
Template "Navigation" 1280x800
   TextField "Template_Text field_1" at 1044,28 size 229x39; Text 'Krauss Maffei'
   Button "Template_Button_17" at 502,23 size 38x32; TextOff 'Text'; PictureOff "Bendera inggris"
      on Click: function_fb9197e8(-1)
   Button "Template_Button_18" at 546,23 size 38x32; TextOff 'Text'; PictureOff "manual mode"
   Button "Template_Button_19" at 590,23 size 38x32; TextOff 'Text'; PictureOff "automatic mode"; PictureList "Operation Mode"
      ProcessValue <- "Operation Mode"
   Button "Template_Button_20" at 634,23 size 38x32; TextOff 'Text'
   Button "Template_Button_21" at 678,23 size 38x32; TextOff 'Text'
   Button "Template_Button_24" at 16,18 size 67x43; TextOff 'Text'; PictureOff "left arrow"
      on Press: function_efd93a16()
   Button "status_reduced" at 678,23 size 38x32; TextOff 'Text'; PictureOff "Reduced green"
      Visibility <- "DB619_State_MPart_Recirculation{1}_Reduced"
   Button "Template_Button_15" at 414,23 size 38x32; TextOff 'Text'
   Button "status_Interval_Reduced" at 678,23 size 38x32; TextOff 'Text'; PictureOff "Interval green"
      Visibility <- "DB619_State_MPart_Recirculation{1}_Intervall_Reduced"
   Button "status_lowpressure" at 678,23 size 38x32; TextOff 'Text'; PictureOff "Lowpress green"
      Visibility <- "DB619_State_MPart_Recirculation{1}_Lowpressure"
   Button "status_Lowpressure_Interval" at 678,23 size 38x32; TextOff 'Text'; PictureOff "lowpress circulation"
      Visibility <- "DB619_State_MPart_Recirculation{1}_Intervall_Lowpressure"
   Button "status_highpressure" at 678,23 size 38x32; TextOff 'Text'; PictureOff "high press circuit"
      Visibility <- "DB619_State_MPart_Recirculation{1}_Highpressure"
   Button "Template_Button_25" at 546,23 size 38x32; TextOff 'Text'; PictureList "Operation Mode"; PictureOff "weekendmode"
      ProcessValue <- "Operation Mode"
      Visibility <- "DB619_State_MPart_Recirculation{1}_Weekendswitching"
   Button "Template_Button_26" at 722,23 size 38x32; TextOff 'Text'
   Button "Template_Button_27" at 678,23 size 38x32; TextOff 'Text'; PictureOff "shot cycle_1"
      Visibility <- "DB619_State_MPart_Cycle{1}_running"
   IOField "Template_I/O field_1" at 97,25 size 273x28; FormatPattern 9999999999999999999999999999999999999999
      ProcessValue <- "TP-Bereichszeiger_Date_Time_ActTime"
   Button "Template_Button_30" at 458,23 size 38x32; TextOff 'Text'
   Button "Template_Button_16" at 458,23 size 38x32; TextOff 'Text'; PictureOff "printer off"; PictureList "Print Function"
      ProcessValue <- "Print Function"
      Visibility <- "Print Function"
   SymbolicIOField "Template_Symbolic I/O field_1" at 800,18 size 120x42; TextOff '0'; TextOn '1'; TextList "MH_NO"
      ProcessValue <- "DB619_State_MPart_SWU{1}_ActualSWU"
   Button "Template_Button_3" at 16,261 size 68x66; TextOff 'Text'; PictureOff "osiloskope"; PictureList "ico_navigation_1"
      on Press: function_b14e0dd5("DB14_TP_Shortcuts_TP_Shortcuts_ButtonNo_2", 0)
      Appearance <- "DB14_TP_Shortcuts_TP_Shortcuts_Page_active_2"
      on Click: ActivateScreenByNumber("DB14_TP_Shortcuts_TP_Shortcuts_PageNo_2", 0)
      Visibility <- "DB14_TP_Shortcuts_TP_Shortcuts_Page_active_2"
      ProcessValue <- "DB14_TP_Shortcuts_TP_Shortcuts_PageNo_2"
   Button "Template_Button_4" at 16,354 size 68x66; TextOff 'Text'; PictureOff "scope_1"; PictureList "ico_navigation_1"
      on Press: function_b14e0dd5("DB14_TP_Shortcuts_TP_Shortcuts_ButtonNo_3", 0)
      on Click: ActivateScreenByNumber("DB14_TP_Shortcuts_TP_Shortcuts_PageNo_3", 0)
      Appearance <- "DB14_TP_Shortcuts_TP_Shortcuts_Page_active_3"
      Visibility <- "DB14_TP_Shortcuts_TP_Shortcuts_Page_active_3"
      ProcessValue <- "DB14_TP_Shortcuts_TP_Shortcuts_PageNo_3"
   Button "Template_Button_6" at 16,539 size 68x66; TextOff 'Text'; PictureOff "s2"; PictureList "ico_navigation_1"
      on Press: function_b14e0dd5("DB14_TP_Shortcuts_TP_Shortcuts_ButtonNo_5", 0)
      on Click: ActivateScreenByNumber("DB14_TP_Shortcuts_TP_Shortcuts_PageNo_5", 0)
      Appearance <- "DB14_TP_Shortcuts_TP_Shortcuts_Page_active_5"
      Visibility <- "DB14_TP_Shortcuts_TP_Shortcuts_Page_active_5"
      ProcessValue <- "DB14_TP_Shortcuts_TP_Shortcuts_PageNo_5"
   Button "Template_Button_13" at 1196,724 size 68x66; TextOff 'Text'; PictureList "Home"; PictureOff "Graphic_8"
      on Click: ActivateScreen("0017_Home Screen", 0)
      Appearance <- "NavScreenChange"
   Button "Template_Button_23" at 1196,631 size 68x66; TextOff 'Text'; PictureList "Nav_Recipe"; PictureOff "chemical"
      on Click: ActivateScreen("0892_Tool Editor", 0)
      Appearance <- "NavScreenChange"
   Button "Template_Button_22" at 1196,446 size 68x66; TextOff 'Text'; PictureOff "archive"; PictureList "Nav_Logging"
      on Click: SetTag("NavScreenChange", 4); SetTag("Recipe_Appearance_Control", 0); SetTag("Archived Alarm Control", 2); SetTag("Archive Alarm Number", 0); "CopyAlarmLogView"(); ActivateScreen("0013_Archive Alarm", 0)
      Appearance <- "NavScreenChange"
   Button "Template_Button_9" at 1196,261 size 68x66; TextOff 'Text'; PictureOff "process"; PictureList "Setting"
      on Click: ActivateScreen("0018_SystemSetting", 0); SetTag("System Setting Screen Control", 0)
      Appearance <- "NavScreenChange"
   Button "Template_Button_2" at 16,169 size 68x66; TextOff 'Text'; PictureList "ico_navigation_1"
      on Press: function_b14e0dd5("DB14_TP_Shortcuts_TP_Shortcuts_ButtonNo_1", 0)
      on Click: ActivateScreenByNumber("DB14_TP_Shortcuts_TP_Shortcuts_PageNo_1", 0)
      Appearance <- "DB14_TP_Shortcuts_TP_Shortcuts_Page_active_1"
      Visibility <- "DB14_TP_Shortcuts_TP_Shortcuts_Page_active_1"
      ProcessValue <- "DB14_TP_Shortcuts_TP_Shortcuts_PageNo_1"
   Button "Template_Button_5" at 16,446 size 68x66; TextOff 'Text'; PictureList "ico_navigation_1"
      on Press: function_b14e0dd5("DB14_TP_Shortcuts_TP_Shortcuts_ButtonNo_4", 0)
      on Click: ActivateScreenByNumber("DB14_TP_Shortcuts_TP_Shortcuts_PageNo_4", 0)
      Appearance <- "DB14_TP_Shortcuts_TP_Shortcuts_Page_active_4"
      Visibility <- "DB14_TP_Shortcuts_TP_Shortcuts_Page_active_4"
      ProcessValue <- "DB14_TP_Shortcuts_TP_Shortcuts_PageNo_4"
   Button "Template_Button_31" at 16,631 size 68x66; TextOff 'Text'; PictureOff "scope_1"; PictureList "ico_navigation_1"
      on Press: function_b14e0dd5("DB14_TP_Shortcuts_TP_Shortcuts_ButtonNo_6", 0)
      on Click: ActivateScreenByNumber("DB14_TP_Shortcuts_TP_Shortcuts_PageNo_6", 0)
      Appearance <- "DB14_TP_Shortcuts_TP_Shortcuts_Page_active_6"
      Visibility <- "DB14_TP_Shortcuts_TP_Shortcuts_Page_active_6"
      ProcessValue <- "DB14_TP_Shortcuts_TP_Shortcuts_PageNo_6"
   Button "Template_Button_7" at 16,724 size 68x66; TextOff 'Text'; PictureList "ico_navigation_1"
      on Press: function_b14e0dd5("DB14_TP_Shortcuts_TP_Shortcuts_ButtonNo_7", 0)
      on Click: ActivateScreenByNumber("DB14_TP_Shortcuts_TP_Shortcuts_PageNo_7", 0)
      Appearance <- "DB14_TP_Shortcuts_TP_Shortcuts_Page_active_7"
      Visibility <- "DB14_TP_Shortcuts_TP_Shortcuts_Page_active_7"
      ProcessValue <- "DB14_TP_Shortcuts_TP_Shortcuts_PageNo_7"
   Button "Template_Button_8" at 1196,169 size 68x66; TextOff 'Text'; PictureOff "Alarm Icon 3"
      on Click: ActivateScreen("0024_ActualFaults", 0); SetTag("NavScreenChange", 1); SetTag("Recipe_Appearance_Control", 0); SetTag("Alarm_Filter_Tag", 0)
      Appearance <- "NavScreenChange"
   Button "Template_Button_10" at 1196,354 size 68x66; TextOff 'Text'
   Button "Template_Button_32" at 1196,539 size 68x66; TextOff 'Text'; PictureOff "049-book"
      on Click: ActivateScreen("0999_Service", 0); SetTag("Service Screen Control Visibility", 0)
      Appearance <- "NavScreenChange"
   Button "Template_Button_11" at 371,23 size 38x32; TextOff 'Text'
      on Click: function_a2a04561()
      Appearance <- "NavUserChange"
   Button "Template_Button_33" at 16,261 size 68x66; TextOff 'Text'; PictureOff "osiloskope"; PictureList "Ico_navigation_2"
      on Click: ActivateScreenByNumber("DB14_TP_Shortcuts_TP_Shortcuts_PageNo_2", 0)
      on Press: function_b14e0dd5("DB14_TP_Shortcuts_TP_Shortcuts_ButtonNo_2", 0)
      Appearance <- "DB14_TP_Shortcuts_TP_Shortcuts_Page_active_2"
      Visibility <- "DB14_TP_Shortcuts_TP_Shortcuts_Page_active_2"
      ProcessValue <- "DB14_TP_Shortcuts_TP_Shortcuts_PageNo_2"
   Button "Template_Button_34" at 16,354 size 68x66; TextOff 'Text'; PictureOff "scope_1"; PictureList "Ico_navigation_2"
      on Press: function_b14e0dd5("DB14_TP_Shortcuts_TP_Shortcuts_ButtonNo_3", 0)
      Appearance <- "DB14_TP_Shortcuts_TP_Shortcuts_Page_active_3"
      Visibility <- "DB14_TP_Shortcuts_TP_Shortcuts_Page_active_3"
      on Click: ActivateScreenByNumber("DB14_TP_Shortcuts_TP_Shortcuts_PageNo_3", 0)
      ProcessValue <- "DB14_TP_Shortcuts_TP_Shortcuts_PageNo_3"
   Button "Template_Button_35" at 16,539 size 68x66; TextOff 'Text'; PictureOff "s2"; PictureList "Ico_navigation_2"
      on Press: function_b14e0dd5("DB14_TP_Shortcuts_TP_Shortcuts_ButtonNo_5", 0)
      Appearance <- "DB14_TP_Shortcuts_TP_Shortcuts_Page_active_5"
      Visibility <- "DB14_TP_Shortcuts_TP_Shortcuts_Page_active_5"
      on Click: ActivateScreenByNumber("DB14_TP_Shortcuts_TP_Shortcuts_PageNo_5", 0)
      ProcessValue <- "DB14_TP_Shortcuts_TP_Shortcuts_PageNo_5"
   Button "Template_Button_36" at 16,169 size 68x66; TextOff 'Text'; PictureList "Ico_navigation_2"
      on Click: ActivateScreenByNumber("DB14_TP_Shortcuts_TP_Shortcuts_PageNo_1", 0)
      on Press: function_b14e0dd5("DB14_TP_Shortcuts_TP_Shortcuts_ButtonNo_1", 0)
      Appearance <- "DB14_TP_Shortcuts_TP_Shortcuts_Page_active_1"
      Visibility <- "DB14_TP_Shortcuts_TP_Shortcuts_Page_active_1"
      ProcessValue <- "DB14_TP_Shortcuts_TP_Shortcuts_PageNo_1"
   Button "Template_Button_37" at 16,446 size 68x66; TextOff 'Text'; PictureList "Ico_navigation_2"
      on Press: function_b14e0dd5("DB14_TP_Shortcuts_TP_Shortcuts_ButtonNo_4", 0)
      Appearance <- "DB14_TP_Shortcuts_TP_Shortcuts_Page_active_4"
      Visibility <- "DB14_TP_Shortcuts_TP_Shortcuts_Page_active_4"
      on Click: ActivateScreenByNumber("DB14_TP_Shortcuts_TP_Shortcuts_PageNo_4", 0)
      ProcessValue <- "DB14_TP_Shortcuts_TP_Shortcuts_PageNo_4"
   Button "Template_Button_38" at 16,631 size 68x66; TextOff 'Text'; PictureOff "scope_1"; PictureList "Ico_navigation_2"
      on Press: function_b14e0dd5("DB14_TP_Shortcuts_TP_Shortcuts_ButtonNo_6", 0)
      Appearance <- "DB14_TP_Shortcuts_TP_Shortcuts_Page_active_6"
      Visibility <- "DB14_TP_Shortcuts_TP_Shortcuts_Page_active_6"
      on Click: ActivateScreenByNumber("DB14_TP_Shortcuts_TP_Shortcuts_PageNo_6", 0)
      ProcessValue <- "DB14_TP_Shortcuts_TP_Shortcuts_PageNo_6"
   Button "Template_Button_39" at 16,724 size 68x66; TextOff 'Text'; PictureList "Ico_navigation_2"
      on Press: function_b14e0dd5("DB14_TP_Shortcuts_TP_Shortcuts_ButtonNo_7", 0)
      Appearance <- "DB14_TP_Shortcuts_TP_Shortcuts_Page_active_7"
      Visibility <- "DB14_TP_Shortcuts_TP_Shortcuts_Page_active_7"
      on Click: ActivateScreenByNumber("DB14_TP_Shortcuts_TP_Shortcuts_PageNo_7", 0)
      ProcessValue <- "DB14_TP_Shortcuts_TP_Shortcuts_PageNo_7"
   Button "Template_Button_40" at 9,160 size 80x636; TextOff 'Text'
      on Click: function_efd93a16("Save", 446, 387, -1, 1, 1)
      Visibility <- "DB_MouldEditor_HMI_uData_sStatusBits"
   Button "Template_Button_47" at 1189,147 size 80x645; TextOff 'Text'
      Visibility <- "DB_MouldEditor_HMI_uData_sStatusBits_xValueChanged"
      on Click: function_efd93a16("Save", 446, 387, -1, -1, 1)
   Button "Template_Button_12" at 9,160 size 80x636; TextOff 'Text'
      on Click: function_efd93a16("Save", 446, 387, -1, -1, 1)
      Visibility <- "DB_MouldEditor_HMI_uData_sStatusBits"
   Button "Template_Button_14" at 1189,147 size 80x645; TextOff 'Text'
      on Click: function_efd93a16("Save", 446, 387, -1, -1, 1)
      Visibility <- "DB_MouldEditor_HMI_uData_sStatusBits_xValueChanged"
      ObjectEnable <- "PopUp_Restrict"
   Button "Template_Button_29" at 9,147 size 80x645; TextOff 'Text'
      on Click: function_efd93a16("Save", 446, 387, -1, -1, 1)
      Visibility <- "DB_MouldEditor_HMI_uData_sStatusBits_xValueChanged"
      ObjectEnable <- "PopUp_Restrict"
   GraphicIOField "Template_Graphic I/O field_1" at 1200,173 size 61x54; PictureList "ico_alarm"
      Visibility <- "DB009_Faults_Fault_State_Grp_1_3_Exist"
      ProcessValue <- "NavScreenChange"
   Button "Template_Button_28" at 1196,167 size 68x66; TextOff 'Text'; PictureOff "Alarm Icon 3"
      on Click: ActivateScreen("0024_ActualFaults", 0); SetTag("Recipe_Appearance_Control", 0); SetTag("Alarm_Filter_Tag", 0)

screen "0021_Machine" 1280x800, template "Navigation"
   on GenerateScreen: SetBit("DB619_State_MPart_Read"); SetTag("Navigation_7", 1)
   TextField "Text field_1" at 426,217 size 232x25; Text 'Autom. runtime interval'
   TextField "Text field_2" at 426,252 size 267x25; Text 'Autom. Break time interval:'
   TextField "Text field_3" at 426,287 size 232x25; Text 'Manual runtime interval'
   TextField "Text field_4" at 426,322 size 260x25; Text 'Manual Break time interval'
   TextField "Text field_6" at 426,392 size 304x25; Text 'Pr.buldup time before 1st shot:'
   TextField "Text field_7" at 426,427 size 176x25; Text 'Flush t. after shot'
   TextField "Text field_8" at 426,462 size 236x25; Text 'Adj. time between shots'
   TextField "Text field_9" at 428,557 size 341x25; Text 'Maximum wait time for shot enable'
   TextField "Text field_10" at 426,592 size 191x25; Text 'Maximum shot time'
   TextField "Text field_11" at 426,627 size 187x25; Text 'Minimum shot time'
   TextField "Text field_12" at 426,662 size 228x25; Text 'Time HP circ. after shot'
   TextField "Text field_15" at 860,217 size 46x25; Text 's'
   TextField "Text field_16" at 860,252 size 46x25; Text 's'
   IOField "autom runtime interval" at 775,213 size 81x32; Authorization "Operate"; FormatPattern 99999
      ProcessValue <- "DB700_Machine_Machine{0}_Int_Runtime_Auto"
   IOField "I/O field_2" at 775,248 size 81x32; Authorization "Operate"; FormatPattern 99999
      ProcessValue <- "DB700_Machine_Machine{0}_Int_Pausetime_Auto"
   IOField "I/O field_3" at 775,283 size 81x32; Authorization "Operate"; FormatPattern 99999
      ProcessValue <- "DB700_Machine_Machine{0}_Int_Runtime_Manual"
   IOField "I/O field_4" at 775,318 size 81x32; Authorization "Operate"; FormatPattern 99999
      ProcessValue <- "DB700_Machine_Machine{0}_Int_Pausetime_Manual"
   IOField "I/O field_6" at 775,388 size 81x32; Authorization "Operate"; FormatPattern 99999
      ProcessValue <- "DB700_Machine_Machine{0}_PressureBuildUpTime"
   IOField "I/O field_7" at 775,423 size 81x32; Authorization "Operate"; FormatPattern 99999
      ProcessValue <- "DB700_Machine_Machine{0}_CtrlChangeTime1"
   IOField "I/O field_8" at 775,458 size 81x32; Authorization "Operate"; FormatPattern 99999
      ProcessValue <- "DB700_Machine_Machine{0}_StandByTime"
   IOField "I/O field_9" at 775,553 size 81x32; Authorization "Operate"; FormatPattern 99999
      ProcessValue <- "DB700_Machine_Machine{0}_Max_WaitTime"
   IOField "I/O field_10" at 775,588 size 81x32; Authorization "Operate"; FormatPattern 99999
      ProcessValue <- "DB700_Machine_Machine{0}_Max_ShotTime"
   IOField "I/O field_11" at 775,623 size 81x32; Authorization "Operate"; FormatPattern 99999
      ProcessValue <- "DB700_Machine_Machine{0}_Min_ShotTime"
   IOField "I/O field_12" at 775,658 size 81x32; Authorization "Operate"; FormatPattern 99999
      ProcessValue <- "DB700_Machine_Machine{0}_HP_time_after_shot"
   TextField "Text field_17" at 860,287 size 46x25; Text 's'
   TextField "Text field_18" at 860,322 size 46x25; Text 's'
   TextField "Text field_20" at 860,392 size 46x25; Text 's'
   TextField "Text field_21" at 860,427 size 46x25; Text 's'
   TextField "Text field_22" at 860,462 size 46x25; Text 's'
   TextField "Text field_23" at 860,557 size 46x25; Text 's'
   TextField "Text field_24" at 860,592 size 46x25; Text 's'
   TextField "Text field_25" at 860,627 size 46x25; Text 's'
   TextField "Text field_26" at 860,662 size 46x25; Text 's'
   Button "Button_3" at 326,104 size 451x32; TextOff 'Machine'
   Button "Button_1" at 392,167 size 513x566; TextOff 'Text'
   Button "Template_Button_41" at 16,724 size 68x66; TextOff 'Text'; PictureList "Ico_navigation_2"; PictureOff "Setting_Nav_7"; Authorization "User administration"
      on Click: ActivateScreen("1000_General Machine Configuration", 0)
      ProcessValue <- "Nav_7"
      Visibility <- "NavUserChange"

screen "0005_Mixinghead Settting" 1280x800, template "Navigation"
   on GenerateScreen: SetBit("DB704_MH_Value_Read"); SetBit("DB614_MH_State_Read"); SetTag("NavScreenChange", 0)
   Button "Button_1" at 125,150 size 519x633; TextOff 'Text'; Authorization "User administration"
   IOField "I/O field_4" at 416,229 size 69x30; Authorization "User administration"; FormatPattern 999
      ProcessValue <- "DB704_MH_Value_Mixinghead{0}_AmountComponent"
   Button "b_Cleaning_Piston" at 424,474 size 45x30; TextOff 'Text'; PictureOff "obeng"
      Visibility <- "DB704_MH_Value_Mixinghead{0}_WithCleaningPiston"
      on Click: SetTag("MH_Control_Visibility", 11)
   Button "b_Interface" at 424,542 size 45x30; TextOff 'Text'; PictureOff "obeng"
      Visibility <- "DB704_MH_Value_Mixinghead{0}_WithInterface"
      on Click: SetTag("MH_Control_Visibility", 12)
   Button "b_Heating" at 424,610 size 45x30; TextOff 'Text'; PictureOff "obeng"
      Visibility <- "DB704_MH_Value_Mixinghead{0}_WithHeating"
      on Click: SetTag("MH_Control_Visibility", 13)
   Button "b_Inerting" at 424,644 size 45x30; TextOff 'Text'; PictureOff "obeng"
      Visibility <- "DB704_MH_Value_Mixinghead{0}_WithInerting"
      on Click: SetTag("MH_Control_Visibility", 14)
   Button "b_Nozzle_Control" at 424,678 size 45x30; TextOff 'Text'; PictureOff "obeng"
      Visibility <- "DB704_MH_Value_Mixinghead{0}_WithNozzleControl"
      on Click: SetTag("MH_Control_Visibility", 15)
   Button "b_Enable_MH" at 424,160 size 45x30; TextOff 'Text'; PictureOff "obeng"
      on Click: SetTag("MH_Control_Visibility", 10)
   IOField "MachineAllocation" at 416,195 size 69x30; Authorization "User administration"; FormatPattern 999
      ProcessValue <- "DB704_MH_Value_Mixinghead{0}_MachineNumber"
   IOField "I/O field_2" at 467,575 size 53x30; Authorization "User administration"; FormatPattern 999
      ProcessValue <- "DB704_MH_Value_Mixinghead{0}_pRrgNumberManual"
   Button "Check_blowing_Device" at 484,745 size 36x32; TextOff 'Text'; PictureList "Check_Uncheck"
      ProcessValue <- "DB704_MH_Value_Mixinghead{0}_WithMHVenting"
      on Click: InvertBit("DB704_MH_Value_Mixinghead{0}_WithMHVenting")
   Button "Check_LowPress" at 484,711 size 36x32; TextOff 'Text'; PictureList "Check_Uncheck"
      ProcessValue <- "DB704_MH_Value_Mixinghead{0}_WithLPCirculation"
      on Click: InvertBit("DB704_MH_Value_Mixinghead{0}_WithLPCirculation")
   Button "Check_Nozzle_Control" at 484,677 size 36x32; TextOff 'Text'; PictureList "Check_Uncheck"
      ProcessValue <- "DB704_MH_Value_Mixinghead{0}_WithNozzleControl"
      on Click: InvertBit("DB704_MH_Value_Mixinghead{0}_WithNozzleControl")
   Button "Check_Inerting" at 484,643 size 36x32; TextOff 'Text'; PictureList "Check_Uncheck"
      ProcessValue <- "DB704_MH_Value_Mixinghead{0}_WithInerting"
      on Click: InvertBit("DB704_MH_Value_Mixinghead{0}_WithInerting")
   Button "Check_Heating" at 484,609 size 36x32; TextOff 'Text'; PictureList "Check_Uncheck"
      ProcessValue <- "DB704_MH_Value_Mixinghead{0}_WithHeating"
      on Click: InvertBit("DB704_MH_Value_Mixinghead{0}_WithHeating")
   Button "Check_Interface" at 484,540 size 36x32; TextOff 'Text'; PictureList "Check_Uncheck"
      ProcessValue <- "DB704_MH_Value_Mixinghead{0}_WithInterface"
      on Click: InvertBit("DB704_MH_Value_Mixinghead{0}_WithInterface")
   Button "Check_99Program" at 484,506 size 36x32; TextOff 'Text'; PictureList "Check_Uncheck"
      ProcessValue <- "DB704_MH_Value_Mixinghead{0}_With99program"
      on Click: InvertBit("DB704_MH_Value_Mixinghead{0}_With99program")
   Button "Check_CleaningPiston" at 484,472 size 36x32; TextOff 'Text'; PictureList "Check_Uncheck"
      ProcessValue <- "DB704_MH_Value_Mixinghead{0}_WithCleaningPiston"
      on Click: InvertBit("DB704_MH_Value_Mixinghead{0}_WithCleaningPiston")
   Button "Check_Enable_MH" at 479,157 size 36x32; TextOff 'Text'; PictureList "Check_Uncheck"
      ProcessValue <- "DB704_MH_Value_Mixinghead{0}_MH_Active"
      on Click: InvertBit("DB704_MH_Value_Mixinghead{0}_MH_Active")
   TextField "Text field_1" at 137,163 size 111x25; Text 'Enable MH:'
   TextField "Text field_2" at 137,197 size 190x25; Text 'Machine allocation:'
   TextField "Text field_3" at 137,231 size 199x25; Text 'Amount Connection:'
   TextField "Text field_4" at 180,269 size 74x25; Text 'No. 01:'
      Visibility <- "DB704_MH_Value_Mixinghead{0}_AmountComponent"
   TextField "Text field_5" at 180,302 size 74x25; Text 'No. 02:'
      Visibility <- "DB704_MH_Value_Mixinghead{0}_AmountComponent"
   TextField "Text field_6" at 137,477 size 171x25; Text 'Cleaning pisteon:'
   TextField "Text field_7" at 137,511 size 122x25; Text '99 Program:'
   TextField "Text field_9" at 137,545 size 100x25; Text 'Interface:'
   TextField "Text field_8" at 137,579 size 178x25; Text 'Start manual prg.:'
   TextField "Text field_10" at 137,613 size 86x25; Text 'Heating:'
   TextField "Text field_14" at 137,749 size 156x25; Text 'Blowing device:'
   TextField "Text field_13" at 137,715 size 139x25; Text 'Low Pressure:'
   TextField "Text field_12" at 137,681 size 151x25; Text 'Nozzle Control:'
   TextField "Text field_11" at 137,647 size 90x25; Text 'Inerting:'
   Button "Button_21" at 819,200 size 216x197; TextOff 'MixingHead'; PictureOff "images_4"
   Button "b_incress_MH_Setting" at 790,104 size 46x32; TextOff 'Text'; PictureOff "right arrow"
      on Click: function_dd21b452("DB614_MH_State_ReadDeviceNo", 1)
   Button "b_decres_MH_Setting" at 267,104 size 46x32; TextOff 'Text'; PictureOff "left arrow"
      on Click: function_b9b71300("DB614_MH_State_ReadDeviceNo", 1)
   Button "Button_3" at 326,104 size 451x32; TextOff 'MH 01'; TextList "MH_NO"
      ProcessValue <- "DB614_MH_State_ReadDeviceNo"
   TextField "Text field_64" at 180,335 size 74x25; Text 'No. 03:'
      Visibility <- "DB704_MH_Value_Mixinghead{0}_AmountComponent"
   TextField "Text field_65" at 180,368 size 74x25; Text 'No. 04:'
      Visibility <- "DB704_MH_Value_Mixinghead{0}_AmountComponent"
   TextField "Text field_66" at 180,401 size 74x25; Text 'No. 05:'
      Visibility <- "DB704_MH_Value_Mixinghead{0}_AmountComponent"
   TextField "Text field_67" at 180,435 size 74x25; Text 'No. 06:'
      Visibility <- "DB704_MH_Value_Mixinghead{0}_AmountComponent"
   SymbolicIOField "Symbolic I/O field_1" at 279,267 size 243x28; TextOff '0'; TextOn '1'; TextList "Pump_Name"
      Visibility <- "DB704_MH_Value_Mixinghead{0}_AmountComponent"
      ProcessValue <- "DB704_MH_Value_Mixinghead{0}_MH_Connection{1}_Pump_No"
   SymbolicIOField "Symbolic I/O field_2" at 279,300 size 243x28; TextOn '1'; TextOff '0'; TextList "Pump_Name"
      Visibility <- "DB704_MH_Value_Mixinghead{0}_AmountComponent"
      ProcessValue <- "DB704_MH_Value_Mixinghead{0}_MH_Connection{2}_Pump_No"
   SymbolicIOField "Symbolic I/O field_3" at 279,333 size 243x28; TextOn '1'; TextOff '0'; TextList "Pump_Name"
      Visibility <- "DB704_MH_Value_Mixinghead{0}_AmountComponent"
      ProcessValue <- "DB704_MH_Value_Mixinghead{0}_MH_Connection{3}_Pump_No"
   SymbolicIOField "Symbolic I/O field_4" at 279,366 size 243x28; TextOn '1'; TextOff '0'; TextList "Pump_Name"
      Visibility <- "DB704_MH_Value_Mixinghead{0}_AmountComponent"
      ProcessValue <- "DB704_MH_Value_Mixinghead{0}_MH_Connection{4}_Pump_No"
   SymbolicIOField "Symbolic I/O field_5" at 279,399 size 243x28; TextOn '1'; TextOff '0'; TextList "Pump_Name"
      Visibility <- "DB704_MH_Value_Mixinghead{0}_AmountComponent"
      ProcessValue <- "DB704_MH_Value_Mixinghead{0}_MH_Connection{5}_Pump_No"
   SymbolicIOField "Symbolic I/O field_6" at 279,432 size 243x28; TextOn '1'; TextOff '0'; TextList "Pump_Name"
      Visibility <- "DB704_MH_Value_Mixinghead{0}_AmountComponent"
      ProcessValue <- "DB704_MH_Value_Mixinghead{0}_MH_Connection{6}_Pump_No"
   Button "Mixinghead_times_trigger" at 1019,259 size 126x89; TextOff 'Times'; PictureOff "Times"
      on Click: SetTag("MH_Control_Visibility", 16)
   Button "Button_14" at 696,528 size 400x222; TextOff 'Text'
      Visibility <- "MH_Control_Visibility"
   IOField "I/O field_5" at 960,680 size 69x30; FormatPattern 99999.999
      Visibility <- "MH_Control_Visibility"
      ProcessValue <- "DB123_MH_IO_Signals_MH{0}_IN_MH_Closingtime"
   Button "Button_26" at 1039,533 size 51x41; TextOff 'Text'; PictureOff "images (1)"
      on Press: SetTag("MH_Control_Visibility", 0)
      Visibility <- "MH_Control_Visibility"
   IOField "I/O field_3" at 960,647 size 69x30; FormatPattern 99999.999
      Visibility <- "MH_Control_Visibility"
      ProcessValue <- "DB123_MH_IO_Signals_MH{0}_IN_MH_Opentime"
   TextField "Text field_15" at 784,560 size 184x25; Text 'Mixing HeadTimes:'
      Visibility <- "MH_Control_Visibility"
   TextField "Text field_16" at 728,613 size 175x25; Text 'General cor. time:'
      Visibility <- "MH_Control_Visibility"
   TextField "Text field_17" at 728,647 size 139x25; Text 'Opening time:'
      Visibility <- "MH_Control_Visibility"
   TextField "Text field_18" at 728,683 size 130x25; Text 'Closing time:'
      Visibility <- "MH_Control_Visibility"
   TextField "Text field_20" at 1030,683 size 46x25; Text 's'
      Visibility <- "MH_Control_Visibility"
   TextField "Text field_56" at 1030,649 size 46x25; Text 's'
      Visibility <- "MH_Control_Visibility"
   IOField "I/O field_14" at 961,611 size 69x30; FormatPattern 99999.999
      Visibility <- "MH_Control_Visibility"
      ProcessValue <- "DB704_MH_Value_Mixinghead{0}_Corrvalue"
   Button "Button_2" at 696,527 size 400x252; TextOff 'Text'
      Visibility <- "MH_Control_Visibility"
   IOField "I/O field_10" at 912,738 size 64x30; FormatPattern 99999
      Visibility <- "MH_Control_Visibility"
      ProcessValue <- "DB704_MH_Value_Mixinghead{0}_DelayTimeNozzlesOff"
   Button "b_Close_MHsetting_NozzleControl" at 1039,532 size 51x41; TextOff 'Text'; PictureOff "images (1)"
      on Press: SetTag("MH_Control_Visibility", 0)
      Visibility <- "MH_Control_Visibility"
   TextField "Text field_22" at 716,538 size 180x29; Text 'Nozzle Control:'
      Visibility <- "MH_Control_Visibility"
   TextField "Text field_23" at 773,588 size 194x25; Text 'with Nozzle/Bypass'
      Visibility <- "MH_Control_Visibility"
   Button "Check_Nozzle_WithNozzle" at 720,584 size 36x32; TextOff 'Text'; PictureList "Check_Uncheck"
      Visibility <- "MH_Control_Visibility"
      on Click: InvertBit("DB704_MH_Value_Mixinghead{0}_WithNozzleControl")
      ProcessValue <- "DB704_MH_Value_Mixinghead{0}_WithNozzleControl"
   Button "Check_Nozzle_Poly" at 720,618 size 36x32; TextOff 'Text'; PictureList "Check_Uncheck"
      Visibility <- "MH_Control_Visibility"
      ProcessValue <- "DB704_MH_Value_Mixinghead{0}_MH_Connection{1}_WithNozzle"
      on Click: InvertBit("DB704_MH_Value_Mixinghead{0}_MH_Connection{1}_WithNozzle")
   Button "Check_Nozzle_Iso" at 927,618 size 36x32; TextOff 'Text'; PictureList "Check_Uncheck"
      Visibility <- "MH_Control_Visibility"
      ProcessValue <- "DB704_MH_Value_Mixinghead{0}_MH_Connection{2}_WithNozzle"
      on Click: InvertBit("DB704_MH_Value_Mixinghead{0}_MH_Connection{2}_WithNozzle")
   Button "Check_Nozzle_Free1" at 720,652 size 36x32; TextOff 'Text'; PictureList "Check_Uncheck"
      Visibility <- "MH_Control_Visibility"
      ProcessValue <- "DB704_MH_Value_Mixinghead{0}_MH_Connection{3}_WithNozzle"
      on Click: InvertBit("DB704_MH_Value_Mixinghead{0}_MH_Connection{3}_WithNozzle")
   Button "Check_Nozzle_Free3" at 927,652 size 36x32; TextOff 'Text'; PictureList "Check_Uncheck"
      Visibility <- "MH_Control_Visibility"
      ProcessValue <- "DB704_MH_Value_Mixinghead{0}_MH_Connection{4}_WithNozzle"
      on Click: InvertBit("DB704_MH_Value_Mixinghead{0}_MH_Connection{4}_WithNozzle")
   Button "Check_Nozzle_Free2" at 720,686 size 36x32; TextOff 'Text'; PictureList "Check_Uncheck"
      Visibility <- "MH_Control_Visibility"
      ProcessValue <- "DB704_MH_Value_Mixinghead{0}_MH_Connection{5}_WithNozzle"
      on Click: InvertBit("DB704_MH_Value_Mixinghead{0}_MH_Connection{5}_WithNozzle")
   Button "Check_Nozzle_Free4" at 927,686 size 36x32; TextOff 'Text'; PictureList "Check_Uncheck"
      Visibility <- "MH_Control_Visibility"
      ProcessValue <- "DB704_MH_Value_Mixinghead{0}_MH_Connection{6}_WithNozzle"
      on Click: InvertBit("DB704_MH_Value_Mixinghead{0}_MH_Connection{6}_WithNozzle")
   TextField "Text field_28" at 720,741 size 160x25; Text 'Switch off delay'
      Visibility <- "MH_Control_Visibility"
   TextField "Text field_29" at 984,741 size 46x25; Text 's'
      Visibility <- "MH_Control_Visibility"
   SymbolicIOField "Symbolic I/O field_7" at 773,623 size 116x22; TextOn '1'; TextOff '0'; TextList "Pump_Name"
      ProcessValue <- "DB704_MH_Value_Mixinghead{0}_MH_Connection{1}_Pump_No"
      Visibility <- "MH_Control_Visibility"
   SymbolicIOField "Symbolic I/O field_8" at 979,623 size 116x22; TextOn '1'; TextOff '0'; TextList "Pump_Name"
      ProcessValue <- "DB704_MH_Value_Mixinghead{0}_MH_Connection{2}_Pump_No"
      Visibility <- "MH_Control_Visibility"
   SymbolicIOField "Symbolic I/O field_9" at 773,657 size 116x22; TextOn '1'; TextOff '0'; TextList "Pump_Name"
      ProcessValue <- "DB704_MH_Value_Mixinghead{0}_MH_Connection{3}_Pump_No"
      Visibility <- "MH_Control_Visibility"
   SymbolicIOField "Symbolic I/O field_10" at 979,657 size 116x22; TextOn '1'; TextOff '0'; TextList "Pump_Name"
      ProcessValue <- "DB704_MH_Value_Mixinghead{0}_MH_Connection{4}_Pump_No"
      Visibility <- "MH_Control_Visibility"
   SymbolicIOField "Symbolic I/O field_11" at 773,691 size 116x22; TextOn '1'; TextOff '0'; TextList "Pump_Name"
      ProcessValue <- "DB704_MH_Value_Mixinghead{0}_MH_Connection{5}_Pump_No"
      Visibility <- "MH_Control_Visibility"
   SymbolicIOField "Symbolic I/O field_12" at 979,691 size 116x22; TextOn '1'; TextOff '0'; TextList "Pump_Name"
      ProcessValue <- "DB704_MH_Value_Mixinghead{0}_MH_Connection{6}_Pump_No"
      Visibility <- "MH_Control_Visibility"
   Button "Button_6" at 695,526 size 400x252; TextOff 'Text'
      Visibility <- "MH_Control_Visibility"
   Button "b_Close_MHSetting_Heating" at 1038,531 size 51x41; TextOff 'Text'; PictureOff "images (1)"
      on Press: SetTag("MH_Control_Visibility", 0)
      Visibility <- "MH_Control_Visibility"
   TextField "Text field_30" at 715,537 size 94x29; Text 'Heating'
      Visibility <- "MH_Control_Visibility"
   TextField "Text field_31" at 766,587 size 114x25; Text 'Mixinghead'
      Visibility <- "MH_Control_Visibility"
   TextField "Text field_32" at 766,621 size 46x25; Text 'Pipe'
      Visibility <- "MH_Control_Visibility"
   TextField "Text field_33" at 766,654 size 59x25; Text 'Spare'
      Visibility <- "MH_Control_Visibility"
   Button "Check_Heating_Mixinghead" at 719,583 size 36x32; TextOff 'Text'; PictureList "Check_Uncheck"
      Visibility <- "MH_Control_Visibility"
      on Click: InvertBit("DB704_MH_Value_Mixinghead{0}_Conf_IntWithMC")
      ProcessValue <- "DB704_MH_Value_Mixinghead{0}_Conf_IntWithMC"
   Button "Check_Heating_Pipe" at 719,617 size 36x32; TextOff 'Text'; PictureList "Check_Uncheck"
      Visibility <- "MH_Control_Visibility"
      on Click: InvertBit("DB704_MH_Value_Mixinghead{0}_Conf_IntWithPlantInerface")
      ProcessValue <- "DB704_MH_Value_Mixinghead{0}_Conf_IntWithPlantInerface"
   Button "Check_Heating_Tubes" at 926,617 size 36x32; TextOff 'Text'; PictureList "Check_Uncheck"
      Visibility <- "MH_Control_Visibility"
      on Click: InvertBit("DB704_MH_Value_Mixinghead{0}_Conf_IntWithCoupler")
      ProcessValue <- "DB704_MH_Value_Mixinghead{0}_Conf_IntWithCoupler"
   TextField "Text field_34" at 971,621 size 61x25; Text 'Tubes'
      Visibility <- "MH_Control_Visibility"
   Button "Check_Heating_Spare1" at 719,650 size 36x32; TextOff 'Text'; PictureList "Check_Uncheck"
      Visibility <- "MH_Control_Visibility"
      on Click: InvertBit("DB704_MH_Value_Mixinghead{0}_Conf_IntWithRobot")
      ProcessValue <- "DB704_MH_Value_Mixinghead{0}_Conf_IntWithRobot"
   Button "Check_Heating_Spare3" at 926,650 size 36x32; TextOff 'Text'; PictureList "Check_Uncheck"
      Visibility <- "MH_Control_Visibility"
      on Click: InvertBit("DB704_MH_Value_Mixinghead{0}_Conf_IntWithMC")
      ProcessValue <- "DB704_MH_Value_Mixinghead{0}_Conf_IntWithMC"
   TextField "Text field_35" at 971,654 size 59x25; Text 'Spare'
      Visibility <- "MH_Control_Visibility"
   TextField "Text field_36" at 766,688 size 59x25; Text 'Spare'
      Visibility <- "MH_Control_Visibility"
   Button "Check_Heating_Spare2" at 719,684 size 36x32; TextOff 'Text'; PictureList "Check_Uncheck"
      Visibility <- "MH_Control_Visibility"
      on Click: InvertBit("DB704_MH_Value_Mixinghead{0}_Conf_IntWithMC")
      ProcessValue <- "DB704_MH_Value_Mixinghead{0}_Conf_IntWithMC"
   Button "Check_Heating_Spare4" at 926,684 size 36x32; TextOff 'Text'; PictureList "Check_Uncheck"
      Visibility <- "MH_Control_Visibility"
      on Click: InvertBit("DB704_MH_Value_Mixinghead{0}_Conf_IntWithMC")
      ProcessValue <- "DB704_MH_Value_Mixinghead{0}_Conf_IntWithMC"
   TextField "Text field_37" at 971,688 size 59x25; Text 'Spare'
      Visibility <- "MH_Control_Visibility"
   Button "Button_12" at 694,525 size 400x252; TextOff 'Text'
      Visibility <- "MH_Control_Visibility"
   Button "b_Close_Interface" at 1037,530 size 51x41; TextOff 'Text'; PictureOff "images (1)"
      Visibility <- "MH_Control_Visibility"
      on Click: SetTag("MH_Control_Visibility", 0)
   TextField "Text field_38" at 714,536 size 120x29; Text 'Interface:'
      Visibility <- "MH_Control_Visibility"
   TextField "Text field_39" at 758,586 size 140x25; Text 'Mould Carrier:'
      Visibility <- "MH_Control_Visibility"
   TextField "Text field_40" at 758,620 size 170x25; Text 'non KM Interface'
      Visibility <- "MH_Control_Visibility"
   TextField "Text field_41" at 758,653 size 62x25; Text 'Robot'
      Visibility <- "MH_Control_Visibility"
   Button "Check_Interface_Mould_Carrier" at 718,582 size 36x32; TextOff 'Text'; PictureList "Check_Uncheck"
      Visibility <- "MH_Control_Visibility"
      on Click: InvertBit("DB704_MH_Value_Mixinghead{0}_Conf_IntWithMC")
      ProcessValue <- "DB704_MH_Value_Mixinghead{0}_Conf_IntWithMC"
   Button "Check_Interface_NonKM" at 718,616 size 36x32; TextOff 'Text'; PictureList "Check_Uncheck"
      Visibility <- "MH_Control_Visibility"
      on Click: InvertBit("DB704_MH_Value_Mixinghead{0}_Conf_IntWithPlantInerface")
      ProcessValue <- "DB704_MH_Value_Mixinghead{0}_Conf_IntWithPlantInerface"
   Button "Check_Interface_DP/DP" at 917,616 size 36x32; TextOff 'Text'; PictureList "Check_Uncheck"
      Visibility <- "MH_Control_Visibility"
      on Click: InvertBit("DB704_MH_Value_Mixinghead{0}_Conf_IntWithCoupler")
      ProcessValue <- "DB704_MH_Value_Mixinghead{0}_Conf_IntWithCoupler"
   TextField "Text field_42" at 957,620 size 147x25; Text 'DP/DP Coupler'
      Visibility <- "MH_Control_Visibility"
   Button "Check_Interface_Robot" at 718,649 size 36x32; TextOff 'Text'; PictureList "Check_Uncheck"
      Visibility <- "MH_Control_Visibility"
      on Click: InvertBit("DB704_MH_Value_Mixinghead{0}_Conf_IntWithRobot")
      ProcessValue <- "DB704_MH_Value_Mixinghead{0}_Conf_IntWithRobot"
   TextField "Text field_44" at 758,687 size 59x25; Text 'Spare'
      Visibility <- "MH_Control_Visibility"
   Button "Check_Interface_Spare" at 718,683 size 36x32; TextOff 'Text'; PictureList "Check_Uncheck"
      Visibility <- "MH_Control_Visibility"
      on Click: InvertBit("DB704_MH_Value_Mixinghead{0}_Conf_IntWithTag")
      ProcessValue <- "DB704_MH_Value_Mixinghead{0}_Conf_IntWithTag"
   Button "Button_16" at 693,524 size 400x252; TextOff 'Text'
      Visibility <- "MH_Control_Visibility"
   Button "bCloseCleanPiston" at 1036,529 size 51x41; TextOff 'Text'; PictureOff "images (1)"
      Visibility <- "MH_Control_Visibility"
      on Click: SetTag("MH_Control_Visibility", 0)
   TextField "Text field_43" at 713,535 size 282x29; Text 'Type of Cleaning Piston:'
      Visibility <- "MH_Control_Visibility"
   TextField "Text field_45" at 777,608 size 81x25; Text 'Interval'
      Visibility <- "MH_Control_Visibility"
   TextField "Text field_46" at 777,642 size 98x25; Text 'Controled'
      Visibility <- "MH_Control_Visibility"
   TextField "Text field_47" at 777,677 size 59x25; Text 'Spare'
      Visibility <- "MH_Control_Visibility"
   Button "Check_CP_Interval" at 717,604 size 36x32; TextOff 'Text'; PictureList "Check_Uncheck"
      Visibility <- "MH_Control_Visibility"
      ProcessValue <- "DB704_MH_Value_Mixinghead{0}_Cleaning_Piston_CP_withInterval"
      on Click: InvertBit("DB704_MH_Value_Mixinghead{0}_Cleaning_Piston_CP_withInterval")
   Button "Check_CP_Controled" at 717,638 size 36x32; TextOff 'Text'; PictureList "Check_Uncheck"
      Visibility <- "MH_Control_Visibility"
      on Click: InvertBit("DB704_MH_Value_Mixinghead{0}_Cleaning_Piston_StepCleaningPiston")
      ProcessValue <- "DB704_MH_Value_Mixinghead{0}_Cleaning_Piston_StepCleaningPiston"
   Button "Check_CP_Regulated" at 924,638 size 36x32; TextOff 'Text'; PictureList "Check_Uncheck"
      Visibility <- "MH_Control_Visibility"
      on Click: InvertBit("DB704_MH_Value_Mixinghead{0}_Cleaning_Piston_ContrCleaningPiston")
      ProcessValue <- "DB704_MH_Value_Mixinghead{0}_Cleaning_Piston_ContrCleaningPiston"
   TextField "Text field_48" at 964,642 size 101x25; Text 'Regulated'
      Visibility <- "MH_Control_Visibility"
   Button "Check_CP_Spare1" at 717,673 size 36x32; TextOff 'Text'; PictureList "Check_Uncheck"
      Visibility <- "MH_Control_Visibility"
      on Click: InvertBit("DB704_MH_Value_Mixinghead{0}_Cleaning_Piston_ContrCleaningPiston")
      ProcessValue <- "DB704_MH_Value_Mixinghead{0}_Cleaning_Piston_ContrCleaningPiston"
   Button "Check_CP_Spare2" at 924,673 size 36x32; TextOff 'Text'; PictureList "Check_Uncheck"
      Visibility <- "MH_Control_Visibility"
      on Click: InvertBit("DB704_MH_Value_Mixinghead{0}_Cleaning_Piston_ContrCleaningPiston")
      ProcessValue <- "DB704_MH_Value_Mixinghead{0}_Cleaning_Piston_ContrCleaningPiston"
   TextField "Text field_49" at 964,677 size 59x25; Text 'Spare'
      Visibility <- "MH_Control_Visibility"
   TextField "Text field_50" at 777,711 size 138x25; Text 'Enable button'
      Visibility <- "MH_Control_Visibility"
   Button "Check_CP_Enable button" at 717,707 size 36x32; TextOff 'Text'; PictureList "Check_Uncheck"
      Visibility <- "MH_Control_Visibility"
      on Click: InvertBit("DB704_MH_Value_Mixinghead{0}_Cleaning_Piston_Spare_19")
      ProcessValue <- "DB704_MH_Value_Mixinghead{0}_Cleaning_Piston_Spare_19"
   Button "Check_CP_Spare3" at 924,707 size 36x32; TextOff 'Text'; PictureList "Check_Uncheck"
      Visibility <- "MH_Control_Visibility"
      on Click: InvertBit("DB704_MH_Value_Mixinghead{0}_Cleaning_Piston_ContrCleaningPiston")
      ProcessValue <- "DB704_MH_Value_Mixinghead{0}_Cleaning_Piston_ContrCleaningPiston"
   TextField "Text field_51" at 964,711 size 59x25; Text 'Spare'
      Visibility <- "MH_Control_Visibility"
   Button "Button_18" at 692,523 size 400x252; TextOff 'Text'
      Visibility <- "MH_Control_Visibility"
   Button "b_Close_MHSetting_MixingType" at 1035,528 size 51x41; TextOff 'Text'; PictureOff "images (1)"
      on Press: SetTag("MH_Control_Visibility", 0)
      Visibility <- "MH_Control_Visibility"
   TextField "Text field_52" at 712,534 size 202x29; Text 'Mixinghead type:'
      Visibility <- "MH_Control_Visibility"
   TextField "Text field_53" at 763,603 size 91x25; Text 'Standard'
      Visibility <- "MH_Control_Visibility"
   TextField "Text field_54" at 763,637 size 71x25; Text 'Analog'
      Visibility <- "MH_Control_Visibility"
   TextField "Text field_55" at 763,671 size 53x25; Text 'Fibre'
      Visibility <- "MH_Control_Visibility"
   Button "Check_MH_Standard" at 716,599 size 36x32; TextOff 'Text'; PictureList "Check_Uncheck"
      Visibility <- "MH_Control_Visibility"
      on Click: InvertBit("DB704_MH_Value_Mixinghead{0}_Conf_MHDigital")
      ProcessValue <- "DB704_MH_Value_Mixinghead{0}_Conf_MHDigital"
   Button "Check_MH_Analog" at 716,633 size 36x32; TextOff 'Text'; PictureList "Check_Uncheck"
      Visibility <- "MH_Control_Visibility"
      on Click: InvertBit("DB704_MH_Value_Mixinghead{0}_Conf_MHControled")
      ProcessValue <- "DB704_MH_Value_Mixinghead{0}_Conf_MHControled"
   Button "Check_MH_Fibre" at 716,667 size 36x32; TextOff 'Text'; PictureList "Check_Uncheck"
      Visibility <- "MH_Control_Visibility"
      on Click: InvertBit("DB704_MH_Value_Mixinghead{0}_Conf_MHFibre")
      ProcessValue <- "DB704_MH_Value_Mixinghead{0}_Conf_MHFibre"
   Button "Check_MH_Spray" at 923,663 size 36x32; TextOff 'Text'; PictureList "Check_Uncheck"
      Visibility <- "MH_Control_Visibility"
      on Click: InvertBit("DB704_MH_Value_Mixinghead{0}_Conf_MHSpray")
      ProcessValue <- "DB704_MH_Value_Mixinghead{0}_Conf_MHSpray"
   TextField "Text field_57" at 969,667 size 59x25; Text 'Spray'
      Visibility <- "MH_Control_Visibility"
   TextField "Text field_58" at 763,705 size 73x25; Text 'Special'
      Visibility <- "MH_Control_Visibility"
   Button "Check_MH_Special" at 716,701 size 36x32; TextOff 'Text'; PictureList "Check_Uncheck"
      Visibility <- "MH_Control_Visibility"
      on Click: InvertBit("DB704_MH_Value_Mixinghead{0}_Conf_MHSpecial")
      ProcessValue <- "DB704_MH_Value_Mixinghead{0}_Conf_MHSpecial"
   Button "Button_22" at 693,523 size 400x252; TextOff 'Text'
      Visibility <- "MH_Control_Visibility"
   Button "b_Close_MHSetting_type" at 1036,528 size 51x41; TextOff 'Text'; PictureOff "images (1)"
      Visibility <- "MH_Control_Visibility"
      on Click: SetTag("MH_Control_Visibility", 0)
   TextField "Text field_59" at 713,534 size 202x29; Text 'Mixinghead type:'
      Visibility <- "MH_Control_Visibility"
   TextField "Text field_60" at 766,603 size 79x25; Text 'OverMH'
      Visibility <- "MH_Control_Visibility"
   TextField "Text field_61" at 770,644 size 71x25; Text 'Analog'
      Visibility <- "MH_Control_Visibility"
   Button "Check_MH_Inerting_OverMH" at 717,599 size 36x32; TextOff 'Text'; PictureList "Check_Uncheck"
      Visibility <- "MH_Control_Visibility"
      on Click: InvertBit("DB704_MH_Value_MH_Inerting{0}_with_inert_over_MH")
      ProcessValue <- "DB704_MH_Value_MH_Inerting{0}_with_inert_over_MH"
   Button "Check_MH_Inerting_Analog" at 717,640 size 36x32; TextOff 'Text'; PictureList "Check_Uncheck"
      Visibility <- "MH_Control_Visibility"
      on Click: InvertBit("DB704_MH_Value_MH_Inerting{0}_with_output_without_N2")
      ProcessValue <- "DB704_MH_Value_MH_Inerting{0}_with_output_without_N2"
   Button "Check_MH_Inerting_Overlance" at 924,599 size 36x32; TextOff 'Text'; PictureList "Check_Uncheck"
      Visibility <- "MH_Control_Visibility"
      on Click: InvertBit("DB704_MH_Value_MH_Inerting{0}_with_inert_over_Lance")
      ProcessValue <- "DB704_MH_Value_MH_Inerting{0}_with_inert_over_Lance"
   TextField "Text field_63" at 972,603 size 103x25; Text 'over lance'
      Visibility <- "MH_Control_Visibility"
   IOField "I/O field_8" at 925,642 size 88x32; FormatPattern 9999.9
      Visibility <- "MH_Control_Visibility"
      ProcessValue <- "DB704_MH_Value_MH_Inerting{0}_Max_Reference_Value_Inert"
   TextField "Text field_62" at 1024,644 size 46x25; Text 'g'
      Visibility <- "MH_Control_Visibility"
   Button "Button_24" at 125,143 size 519x643; TextOff 'Text'; Authorization "User administration"; PictureOff "images_4"
      Visibility <- "DB704_MH_Value_Mixinghead{0}_MH_Active"
      on Press: SetBit("DB704_MH_Value_Mixinghead{0}_MH_Active")

